REGION Network 26: Head status
   RUNG wire#powerrail
      Contact( "AlwaysTRUE" )
      wire#w1
      I_Contact( #OUTPUT_xFireON )
      Move(in := 1, out1 => #tHMR.dHeadStatus)
   END_RUNG
   RUNG wire#w1
      Contact( #OUTPUT_xFireON )
      Move(in := 3, out1 => #tHMR.dHeadStatus)
   END_RUNG
   // the same network as SCL:
   IF "AlwaysTRUE" AND NOT #OUTPUT_xFireON THEN #tHMR.dHeadStatus := 1; END_IF;
   IF "AlwaysTRUE" AND #OUTPUT_xFireON THEN #tHMR.dHeadStatus := 3; END_IF;
END_REGION

REGION Network 27: Head#x reset head usage counter {x|x|x|x|O}
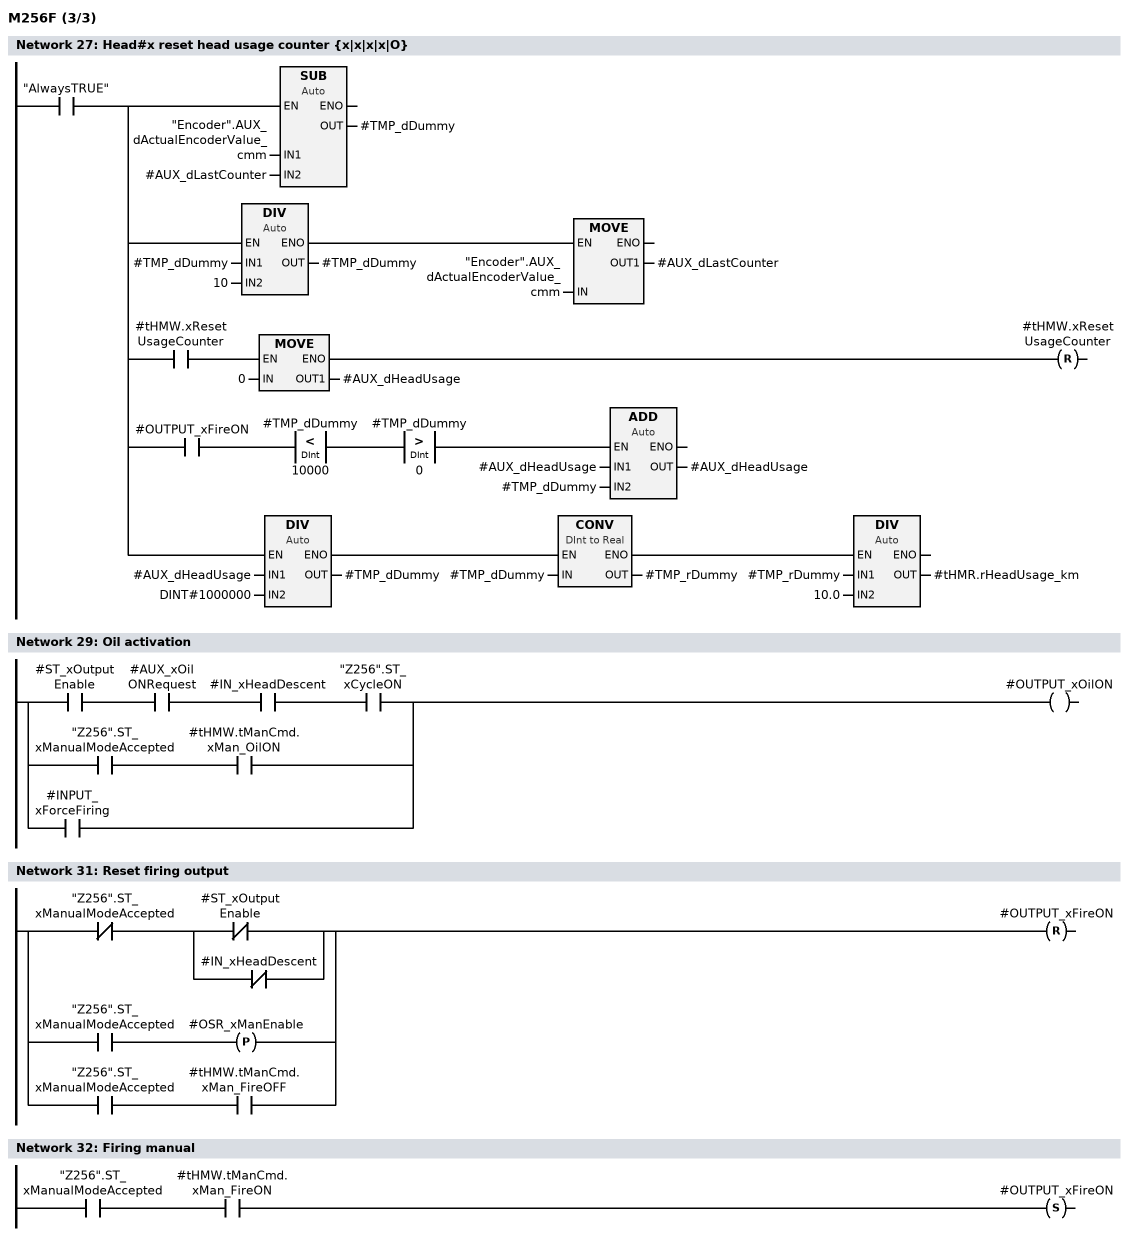
   RUNG wire#powerrail
      Contact( "AlwaysTRUE" )
      wire#w1
      Sub(in1 := "Encoder".AUX_dActualEncoderValue_cmm, in2 := #AUX_dLastCounter, out => #TMP_dDummy)
   END_RUNG
   RUNG wire#w1
      Div(in1 := #TMP_dDummy, in2 := 10, out => #TMP_dDummy)
      Move(in := "Encoder".AUX_dActualEncoderValue_cmm, out1 => #AUX_dLastCounter)
   END_RUNG
   RUNG wire#w1
      Contact( #tHMW.xResetUsageCounter )
      Move(in := 0, out1 => #AUX_dHeadUsage)
      R_Coil( #tHMW.xResetUsageCounter )
   END_RUNG
   RUNG wire#w1
      Contact( #OUTPUT_xFireON )
      { S7_Templates := "SrcType := DInt" } LT_Contact(in1 := #TMP_dDummy, in2 := 10000)
      { S7_Templates := "SrcType := DInt" } GT_Contact(in1 := #TMP_dDummy, in2 := 0)
      Add(in1 := #AUX_dHeadUsage, in2 := #TMP_dDummy, out => #AUX_dHeadUsage)
   END_RUNG
   RUNG wire#w1
      Div(in1 := #AUX_dHeadUsage, in2 := DINT#1000000, out => #TMP_dDummy)
      { S7_Templates := "[SrcType := DInt, DestType := Real]" } Convert(in := #TMP_dDummy, out => #TMP_rDummy)
      Div(in1 := #TMP_rDummy, in2 := 10.0, out => #tHMR.rHeadUsage_km)
   END_RUNG
   // the same network as SCL:
   IF "AlwaysTRUE" THEN
       #TMP_dDummy := "Encoder".AUX_dActualEncoderValue_cmm - #AUX_dLastCounter;
       #TMP_dDummy := #TMP_dDummy / 10;
       #AUX_dLastCounter := "Encoder".AUX_dActualEncoderValue_cmm;
   END_IF;
   IF "AlwaysTRUE" AND #tHMW.xResetUsageCounter THEN
       #AUX_dHeadUsage := 0;
       #tHMW.xResetUsageCounter := FALSE;
   END_IF;
   IF "AlwaysTRUE" AND #OUTPUT_xFireON AND (#TMP_dDummy < 10000) AND (#TMP_dDummy > 0) THEN
       #AUX_dHeadUsage := #AUX_dHeadUsage + #TMP_dDummy;
   END_IF;
   IF "AlwaysTRUE" THEN
       #TMP_dDummy := #AUX_dHeadUsage / DINT#1000000;
       #TMP_rDummy := DINT_TO_REAL(#TMP_dDummy);
       #tHMR.rHeadUsage_km := #TMP_rDummy / 10.0;
   END_IF;
END_REGION

REGION Network 28: ####_OUTPUT_####
END_REGION

REGION Network 29: Oil activation
   RUNG wire#powerrail
      Contact( #ST_xOutputEnable )
      Contact( #AUX_xOilONRequest )
      Contact( #IN_xHeadDescent )
      Contact( "Z256".ST_xCycleON )
      wire#w1
      Coil( #OUTPUT_xOilON )
   END_RUNG
   RUNG wire#powerrail
      Contact( "Z256".ST_xManualModeAccepted )
      Contact( #tHMW.tManCmd.xMan_OilON )
   END_RUNG wire#w1
   RUNG wire#powerrail
      Contact( #INPUT_xForceFiring )
   END_RUNG wire#w1
   // the same network as SCL:
   #OUTPUT_xOilON := (#ST_xOutputEnable AND #AUX_xOilONRequest AND #IN_xHeadDescent AND "Z256".ST_xCycleON) OR ("Z256".ST_xManualModeAccepted AND #tHMW.tManCmd.xMan_OilON) OR #INPUT_xForceFiring;
END_REGION

REGION Network 30 (SCL): Pressure to heads and display
   #TMP_rDummy := DINT_TO_REAL("CONST_dPressureMax_Unit"-"CONST_dPressureMin_Unit")/ DINT_TO_REAL("CONST_dPressureMax_MN"-"CONST_dPressureMin_MN");
   #TMP_dDummy :=#tHMW.dHeadPressure_mN-"CONST_dPressureMin_MN";
   #OUTPUT_iPressuremA := REAL_TO_INT(#TMP_rDummy *  DINT_TO_REAL(#TMP_dDummy))+DINT_TO_INT("CONST_dPressureMin_Unit");

   IF "CM_IDEV_FromMainLine".xQLTplate THEN
       #OUTPUT_iPressuremA := #OUTPUT_iPressuremA / 100 * DINT_TO_INT("Z256_hmi".tHMW.dPressureScalerOnSample_perc);
   END_IF;
END_REGION

REGION Network 31: Reset firing output
   RUNG wire#powerrail
      I_Contact( "Z256".ST_xManualModeAccepted )
      wire#w1
      I_Contact( #ST_xOutputEnable )
      wire#w2
      R_Coil( #OUTPUT_xFireON )
   END_RUNG
   RUNG wire#w1
      I_Contact( #IN_xHeadDescent )
   END_RUNG wire#w2
   RUNG wire#powerrail
      Contact( "Z256".ST_xManualModeAccepted )
      P_Trig( #OSR_xManEnable )
   END_RUNG wire#w2
   RUNG wire#powerrail
      Contact( "Z256".ST_xManualModeAccepted )
      Contact( #tHMW.tManCmd.xMan_FireOFF )
   END_RUNG wire#w2
   // the same network as SCL:
   #_w1 := "Z256".ST_xManualModeAccepted AND NOT #OSR_xManEnable;   // rising edge
   #OSR_xManEnable := "Z256".ST_xManualModeAccepted;
   IF (NOT "Z256".ST_xManualModeAccepted AND (NOT #ST_xOutputEnable OR NOT #IN_xHeadDescent)) OR #_w1 OR ("Z256".ST_xManualModeAccepted AND #tHMW.tManCmd.xMan_FireOFF) THEN
       #OUTPUT_xFireON := FALSE;
   END_IF;
END_REGION

REGION Network 32: Firing manual
   RUNG wire#powerrail
      Contact( "Z256".ST_xManualModeAccepted )
      Contact( #tHMW.tManCmd.xMan_FireON )
      S_Coil( #OUTPUT_xFireON )
   END_RUNG
   // the same network as SCL:
   IF "Z256".ST_xManualModeAccepted AND #tHMW.tManCmd.xMan_FireON THEN #OUTPUT_xFireON := TRUE; END_IF;
END_REGION
END_FUNCTION_BLOCK

FUNCTION_BLOCK "M256M"   // FB101, LAD
{ S7_Optimized_Access := 'TRUE' }
VERSION : 0.1
   VAR_INPUT
      IN_tConnectionData : "UDT_MB_ConnData";   // IP and connection ID
      IN_dHeadCycleIndex : DInt;   // Number of head cycle (Actual head-1)
      IN_xST_AllHeadStoppingFaults : Bool;   // Cumulative head alarm
      IN_ST_xAllHeadInitialized : Bool;   // All head initialized
      IN_ST_xAllHeadPositioned : Bool;   // All head positioned
      IN_ST_xAllHeadReferred : Bool;   // All head referred
   END_VAR
   VAR
      ST_xHeadInitialized : Bool;   // Head #x initialized
      ST_xHeadReferredSwitch : Bool;   // Head #x referred
      ST_xHeadPositioned : Bool;   // Head #x positioned
      ST_xOutputEnable : Bool;   // Head #x output enable
      ST_xPhaseInProgress : Bool;   // Head #x phases in progress
      ST_xStoppingFaults : Bool;   // Head #x in stopping fault
      ST_xWarnings : Bool;   // Head #x in warning
      ST_xMovementInProgress : Bool;   // Head #x in movement
      ST_xFaults : Bool;   // Head #x in faults
      ST_xHeadVirtualCollision : Bool;   // Head #x virtual collision
      ST_xHeadIPAvail : Bool;   // Head #x is IP linked
      ST_xBrakeReleaseRequest : Bool;   // Head #x brake release requested
      ST_xConditionOKforPowerON : Bool;   // Head #x power on condition
      OSR_xAllHeadReferred : Bool;   // OSR all hed referred
      OSR_xDriveEnable : Bool;   // OSR drive enable
      OSR_xBrakeReleaseSB : Bool;   // OS Brake release
      OS_xBrakeReleaseSB : Bool;   // OS Brake release
      OS_xBrakeRelease : Bool;   // OS Brake release
      OS_xBrakeEngage : Bool;   // OS Brake engaged
      ON_xMotorMBReset : Bool;   // ON Modbus motor reset
      OSN_xMotorMBReset : Bool;   // OSN Modbus motor reset
      INPUT_xOverstroke : Bool;   // Head #x Carriage overstroke
      INPUT_xBrakeRelease : Bool;   // Head #x Brake release button
      INPUT_xCarriageOverload : Bool;   // Head #x Carriage overload
      PH_xHeadInit : Bool;   // Head #x initialization in progress
      PH_xHeadEndInit : Bool;   // Head #x end initialization in progress
      PH_xHeadHomeSwitch : Bool;   // Head #x home in progress to switch
      PH_xHeadEndHomeSwitch : Bool;   // Head #x end home in progress to switch
      PH_xHeadPositioning : Bool;   // Head #x positioning in progress
      PH_xHeadEndPositioning : Bool;   // Head #x end positioning in progress
      AUX_tModbusTCP : TCP_MB_FC8_Req;   // Modbus data
      AUX_xPosCadencer : Bool;   // Cadencer head #x - Positioning allowed
      AUX_dHeadRequestPosition_cmm : DInt;   // Head #x request position [mm/100]
      AUX_dHeadActualPosition_cmm : DInt;   // Head #x actual position [mm/100]
      AUX_rDistanceSwitchTo0 : Real;   // Head #x distance 0 encoder to cam
      AUX_dHeadActSpeed : DInt;   // Head #x actual speed
      AUX_dActualDownloadPar : DInt;   // Head #x actual parameter in download
      AUX_xHomeCadencer : Bool;   // Cadencer head #x - Home position allowed
      AUX_tmDriveReadyRetainTimer : IEC_TIMER;   // Drive ready retain timer
      AUX_tmHeadPositioningTimeout : IEC_TIMER;   // Positioning timeout timer
      AUX_tmHeadHomingTimeout : IEC_TIMER;   // Homing timeout timer
      AUX_tmOFFComOK : IEC_TIMER;   // Head communication OK retained
      AUX_tmOFFEnablePositioningAfterHome : IEC_TIMER;   // Wait drive positioning after homing
      AUX_tmOFFDriveEnable : IEC_TIMER;   // Wait drive enable
      AUX_tmOFFReadCamOffsetAfterHome : IEC_TIMER;   // Retained read cam offset after homing
      AUX_tmHeadInitTimeout : IEC_TIMER;   // Initialization timeout timer
      Axis_Ref : "ILx2T_Ref";
      ILx2_ModbusTCP_Data_Instance : "ILx2_ModbusTCP_Data_1500";
      ILx2T_Control_Instance : "ILx2T_Control";
      ILx2T_Homing_Instance : "ILx2T_Homing";
      ILx2T_Jog_Instance : "ILx2T_Jog";
      ILx2T_ProfilePosition_Instance : "ILx2T_ProfilePosition";
      ILx2T_ProfileVelocity_Instance : "ILx2T_ProfileVelocity";
      ILx2T_Parameter_Read_Write_Instance_Pos : "ILx2T_Parameter_Read_Write";
      ILx2T_Parameter_Read_Write_Instance_Cam : "ILx2T_Parameter_Read_Write";
      ILx2T_Parameter_Read_Write_Instance_Speed : "ILx2T_Parameter_Read_Write";
      ILx2T_Parameter_Read_Write_Instance : "ILx2T_Parameter_Read_Write";
   END_VAR
   VAR RETAIN
      tHMR : Struct   // {[Unit][Scada unit][Low limit][High limit][Access]}
         iCodeAlarm : Int;
         dHeadActualPositions_cmm : DInt;   // Head#x head actual position [mm/100] {mm/100|mm|x|x|O} / Head #x head actual position [mm/100] {mm/100|mm|x|x|O}
         dHeadHomePositions_cmm : DInt;   // Head#x home position [mm/100] {mm/100|mm|x|x|O} / Head #x home position [mm/100] {mm/100|mm|x|x|O}
         rgdHeadMoveStatus : DInt;   // Head#x move status (1=Not Initialized 2=Not referred 3=Not positioned 4=Positioned 5=Positioning 6=Virtual collision 7=Anomaly) {x|x|x|x|O} / Head #x move status (1=Not Initialized 2=Not referred 3=Not positioned 4=Positioned 5=Positioning 6=Virtual collision 7=Anomaly) {x|x|x|x|O}
         tManCmd : Struct
            xMan_JogForwardFdbk : Bool;   // Head#x manual jog forward fdbk {x|x|x|x|O} / Head #x manual jog forward fdbk {x|x|x|x|O}
            xMan_JogBackwardFdbk : Bool;   // Head#x manual jog backward fdbk {x|x|x|x|O} / Head #x manual jog backward fdbk {x|x|x|x|O}
         END_STRUCT;
      END_STRUCT;
      tHMW : Struct   // {[Unit][Scada unit][Low limit][High limit][Access]}
         xBrakeRealeaseHeads : Bool := FALSE;   // Force the brake release of the head {x|x|x|x|M}
         xBrakeEngageHeads : Bool := FALSE;   // Force the brake engaged of the head {x|x|x|x|M}
         xUpdateHomeHead : Bool;   // Update home position head#x {x|x|x|x|M} / Update home position Head #x {x|x|x|x|M}
         dHeadHomePositions_cmm : DInt;   // Head#x home position [mm/100] {mm/100|mm|-2500|2500|M} / Head #x home position [mm/100] {mm/100|mm|-2500|2500|M}
         tManCmd : Struct
            xMan_JogBackward : Bool;   // Head #x manual jog backward {x|x|x|x|O}
            xMan_JogForward : Bool;   // Head #x manual jog forward {x|x|x|x|O}
         END_STRUCT;
      END_STRUCT;
   END_VAR
   VAR
      tALM : Struct
         tW : Struct
            x0 : Bool;
            x1 : Bool;
            x2 : Bool;
            x3 : Bool;
            x4 : Bool;
            x5 : Bool;
            x6 : Bool;
            x7 : Bool;
            x8 : Bool;
            x9 : Bool;
            x10 : Bool;
            x11 : Bool;
            x12 : Bool;
            x13 : Bool;
            x14 : Bool;
            x15 : Bool;
            x16 : Bool;
            x17 : Bool;
            x18 : Bool;
            x19 : Bool;
            x20 : Bool;
            x21 : Bool;
            x22 : Bool;
            x23 : Bool;
            x24 : Bool;
            x25 : Bool;
            x26 : Bool;
            x27 : Bool;
            x28 : Bool;
            x29 : Bool;
            x30 : Bool;
            x31 : Bool;
         END_STRUCT;
         tS : Struct
            x0 : Bool;   // Head#x Initialization timeout / Head #x Initialization timeout
            x1 : Bool;   // Head#x homing timeout / Head #x homing timeout
            x2 : Bool;   // Head#x positioning timeout / Head #x positioning timeout
            x3 : Bool;   // Head#x carriage overload / Head #x carriage overload
            x4 : Bool;   // Head#x drive error / Head #x drive error
            x5 : Bool;   // Head#x missing ethernet IP connection / Head #x missing ethernet IP connection
            x6 : Bool;   // Head op.side overstroke
            x7 : Bool;   // Head oppo.op.side overstroke
            x8 : Bool;   // Head #x overstroke
            x9 : Bool;
            x10 : Bool;
            x11 : Bool;
            x12 : Bool;
            x13 : Bool;
            x14 : Bool;
            x15 : Bool;
            x16 : Bool;
            x17 : Bool;
            x18 : Bool;
            x19 : Bool;
            x20 : Bool;
            x21 : Bool;
            x22 : Bool;
            x23 : Bool;
            x24 : Bool;
            x25 : Bool;
            x26 : Bool;
            x27 : Bool;
            x28 : Bool;
            x29 : Bool;
            x30 : Bool;
            x31 : Bool;
         END_STRUCT;
         tF : Struct
            x0 : Bool;
            x1 : Bool;
            x2 : Bool;
            x3 : Bool;
            x4 : Bool;
            x5 : Bool;
            x6 : Bool;
            x7 : Bool;
            x8 : Bool;
            x9 : Bool;
            x10 : Bool;
            x11 : Bool;
            x12 : Bool;
            x13 : Bool;
            x14 : Bool;
            x15 : Bool;
            x16 : Bool;
            x17 : Bool;
            x18 : Bool;
            x19 : Bool;
            x20 : Bool;
            x21 : Bool;
            x22 : Bool;
            x23 : Bool;
            x24 : Bool;
            x25 : Bool;
            x26 : Bool;
            x27 : Bool;
            x28 : Bool;
            x29 : Bool;
            x30 : Bool;
            x31 : Bool;
         END_STRUCT;
      END_STRUCT;
   END_VAR
   VAR_TEMP
      TMP_rDummy : Real;
      TMP_dwDummy : DWord;
      TMP_dDummy : DInt;
      TMP_dPosition : DInt;
      TMP_dIndex2Nd : DInt;
      TMP_xWriteDoneOS : Bool;
      TMP_xRead : Bool;
      TMP_xMotorOFF : Bool;
   END_VAR
   VAR_TEMP   // added for the SCL form of the ladder/FBD networks
      _w1 : Bool;
      _w2 : Bool;
   END_VAR
   // ILx2T_Homing_Instance.i_diHMsrchdisusr := 0;
BEGIN

REGION Network 1: ####_COSTANTS_####
END_REGION

REGION Network 2: ####_ALARMS_####
END_REGION

REGION Network 3: Reset faults
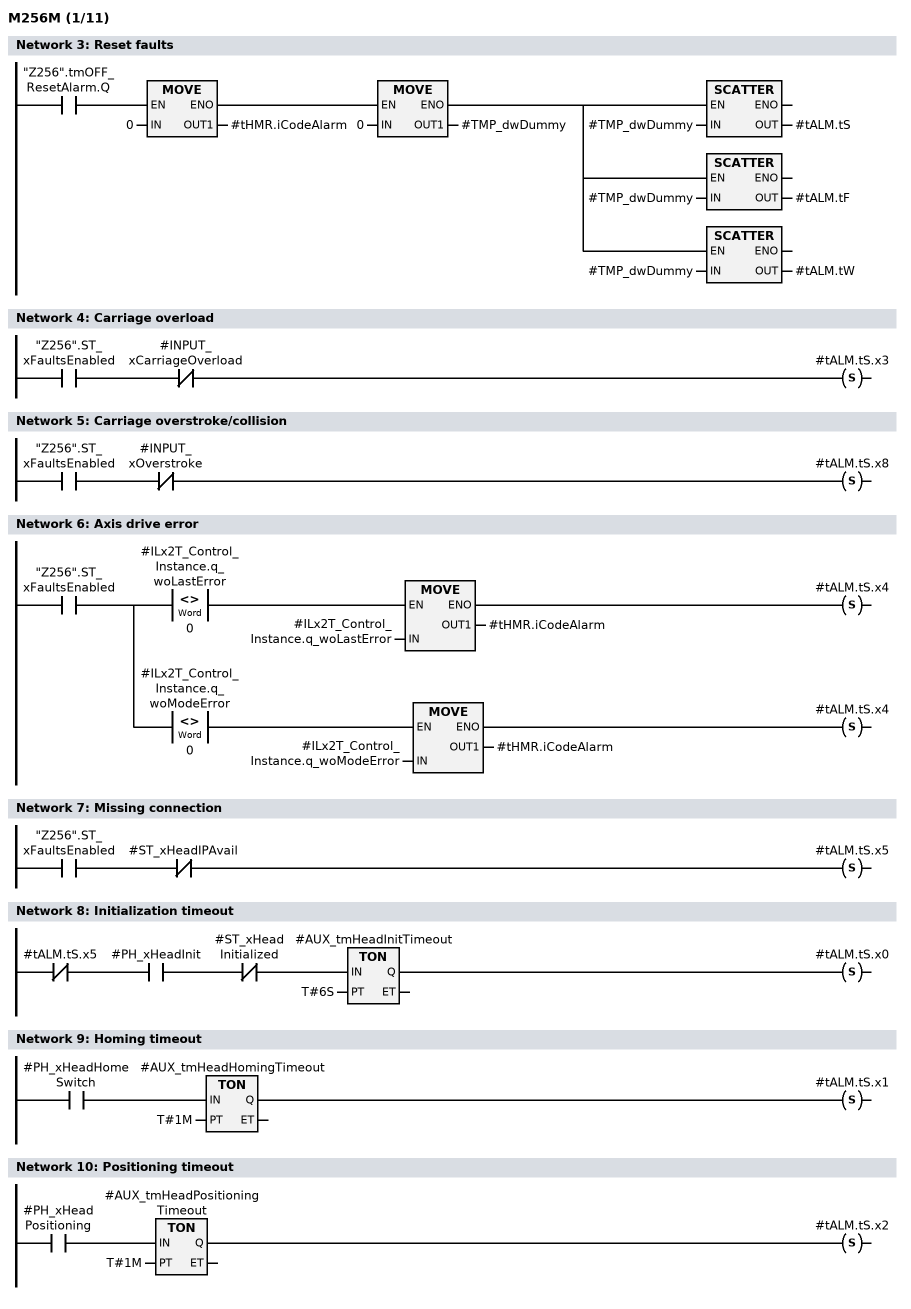
   IF "Z256".tmOFF_ResetAlarm.Q THEN
       #tHMR.iCodeAlarm := 0;
       #TMP_dwDummy := 0;
   END_IF;
   #_w1 := "Z256".tmOFF_ResetAlarm.Q;
   IF #_w1 THEN
       SCATTER(IN := #TMP_dwDummy, OUT => #tALM.tS);
       SCATTER(IN := #TMP_dwDummy, OUT => #tALM.tF);
       SCATTER(IN := #TMP_dwDummy, OUT => #tALM.tW);
   END_IF;
END_REGION

REGION Network 4: Carriage overload
   RUNG wire#powerrail
      Contact( "Z256".ST_xFaultsEnabled )
      I_Contact( #INPUT_xCarriageOverload )
      S_Coil( #tALM.tS.x3 )
   END_RUNG
   // the same network as SCL:
   IF "Z256".ST_xFaultsEnabled AND NOT #INPUT_xCarriageOverload THEN #tALM.tS.x3 := TRUE; END_IF;
END_REGION

REGION Network 5: Carriage overstroke/collision
   RUNG wire#powerrail
      Contact( "Z256".ST_xFaultsEnabled )
      I_Contact( #INPUT_xOverstroke )
      S_Coil( #tALM.tS.x8 )
   END_RUNG
   // the same network as SCL:
   IF "Z256".ST_xFaultsEnabled AND NOT #INPUT_xOverstroke THEN #tALM.tS.x8 := TRUE; END_IF;
END_REGION

REGION Network 6: Axis drive error
   RUNG wire#powerrail
      Contact( "Z256".ST_xFaultsEnabled )
      wire#w1
      { S7_Templates := "SrcType := Word" } NE_Contact(in1 := #ILx2T_Control_Instance.q_woLastError, in2 := 0)
      Move(in := #ILx2T_Control_Instance.q_woLastError, out1 => #tHMR.iCodeAlarm)
      S_Coil( #tALM.tS.x4 )
   END_RUNG
   RUNG wire#w1
      { S7_Templates := "SrcType := Word" } NE_Contact(in1 := #ILx2T_Control_Instance.q_woModeError, in2 := 0)
      Move(in := #ILx2T_Control_Instance.q_woModeError, out1 => #tHMR.iCodeAlarm)
      S_Coil( #tALM.tS.x4 )
   END_RUNG
   // the same network as SCL:
   IF "Z256".ST_xFaultsEnabled AND (#ILx2T_Control_Instance.q_woLastError <> 0) THEN
       #tHMR.iCodeAlarm := #ILx2T_Control_Instance.q_woLastError;
       #tALM.tS.x4 := TRUE;
   END_IF;
   IF "Z256".ST_xFaultsEnabled AND (#ILx2T_Control_Instance.q_woModeError <> 0) THEN
       #tHMR.iCodeAlarm := #ILx2T_Control_Instance.q_woModeError;
       #tALM.tS.x4 := TRUE;
   END_IF;
END_REGION

REGION Network 7: Missing connection
   RUNG wire#powerrail
      Contact( "Z256".ST_xFaultsEnabled )
      I_Contact( #ST_xHeadIPAvail )
      S_Coil( #tALM.tS.x5 )
   END_RUNG
   // the same network as SCL:
   IF "Z256".ST_xFaultsEnabled AND NOT #ST_xHeadIPAvail THEN #tALM.tS.x5 := TRUE; END_IF;
END_REGION

REGION Network 8: Initialization timeout
   #AUX_tmHeadInitTimeout.TON(IN := NOT #tALM.tS.x5 AND #PH_xHeadInit AND NOT #ST_xHeadInitialized, PT := T#6S);
   IF #AUX_tmHeadInitTimeout.Q THEN #tALM.tS.x0 := TRUE; END_IF;
END_REGION

REGION Network 9: Homing timeout
   #AUX_tmHeadHomingTimeout.TON(IN := #PH_xHeadHomeSwitch, PT := T#1M);
   IF #AUX_tmHeadHomingTimeout.Q THEN #tALM.tS.x1 := TRUE; END_IF;
END_REGION

REGION Network 10: Positioning timeout
   #AUX_tmHeadPositioningTimeout.TON(IN := #PH_xHeadPositioning, PT := T#1M);
   IF #AUX_tmHeadPositioningTimeout.Q THEN #tALM.tS.x2 := TRUE; END_IF;
END_REGION

REGION Network 11 (SCL): Cumulative of warning active
   #ST_xWarnings := 0;

   GATHER(IN:= #tALM.tW,
          OUT=>#TMP_dwDummy);

   IF #TMP_dwDummy <> 0 THEN
       #ST_xWarnings := 1;
   END_IF;
END_REGION

REGION Network 12 (SCL): Cumulative of stopping faults active
   #ST_xStoppingFaults := 0;
   GATHER(IN := #tALM.tS,
          OUT => #TMP_dwDummy);

   IF #TMP_dwDummy <> 0 THEN
       #ST_xStoppingFaults := 1;
   END_IF;
END_REGION

REGION Network 13 (SCL): Cumulative of faults active
   #ST_xFaults := 0;
   GATHER(IN := #tALM.tF,
          OUT => #TMP_dwDummy);

   IF #TMP_dwDummy <> 0 THEN
       #ST_xFaults := 1;
   END_IF;
END_REGION

REGION Network 14: #####_HMI LOGICS_#####
END_REGION

REGION Network 15: OS Brake release
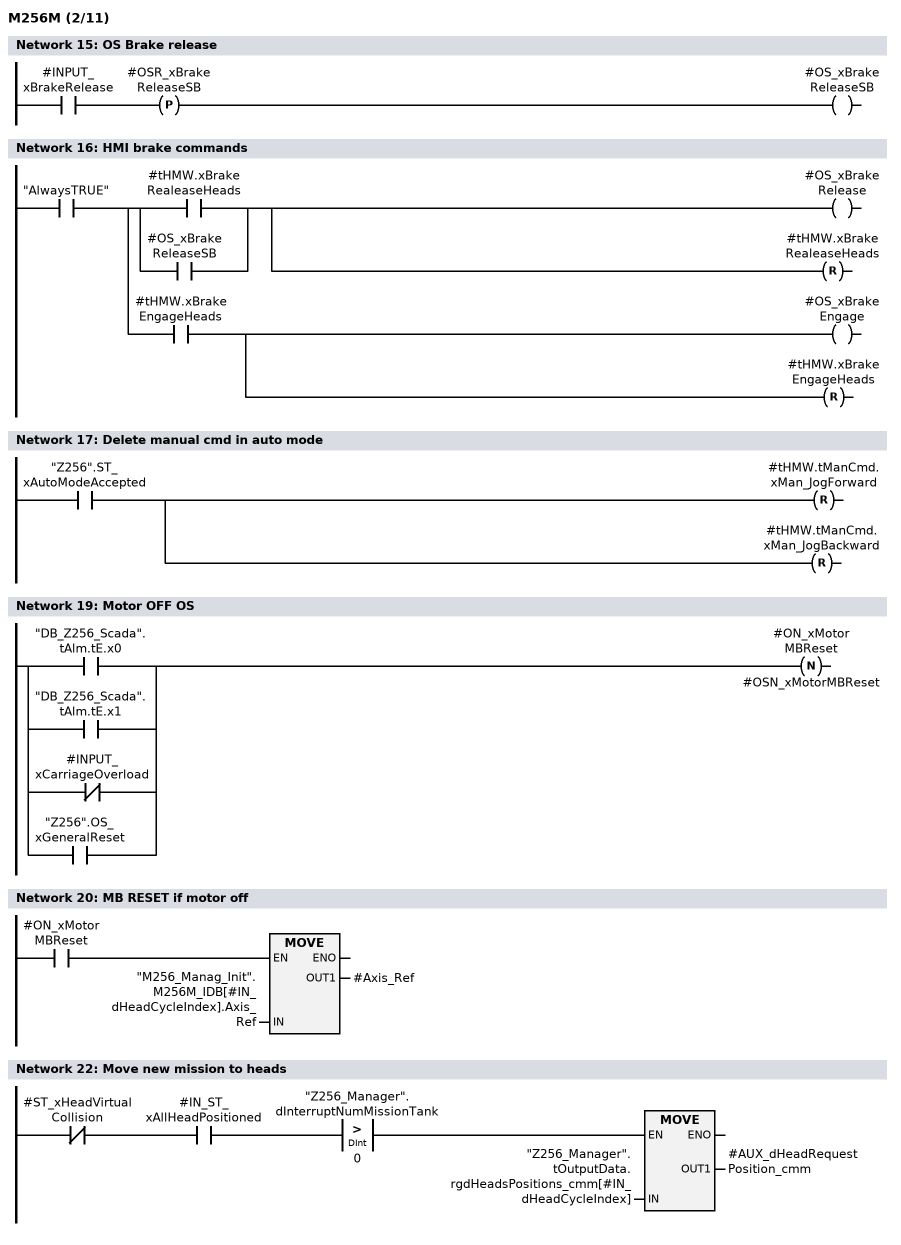
   RUNG wire#powerrail
      Contact( #INPUT_xBrakeRelease )
      P_Trig( #OSR_xBrakeReleaseSB )
      Coil( #OS_xBrakeReleaseSB )
   END_RUNG
   // the same network as SCL:
   #_w1 := #INPUT_xBrakeRelease AND NOT #OSR_xBrakeReleaseSB;   // rising edge
   #OSR_xBrakeReleaseSB := #INPUT_xBrakeRelease;
   #OS_xBrakeReleaseSB := #_w1;
END_REGION

REGION Network 16: HMI brake commands
   RUNG wire#powerrail
      Contact( "AlwaysTRUE" )
      wire#w1
      Contact( #tHMW.xBrakeRealeaseHeads )
      wire#w2
      Coil( #OS_xBrakeRelease )
   END_RUNG
   RUNG wire#w1
      Contact( #OS_xBrakeReleaseSB )
   END_RUNG wire#w2
   RUNG wire#w2
      R_Coil( #tHMW.xBrakeRealeaseHeads )
   END_RUNG
   RUNG wire#w1
      Contact( #tHMW.xBrakeEngageHeads )
      wire#w3
      Coil( #OS_xBrakeEngage )
   END_RUNG
   RUNG wire#w3
      R_Coil( #tHMW.xBrakeEngageHeads )
   END_RUNG
   // the same network as SCL:
   #OS_xBrakeRelease := "AlwaysTRUE" AND (#tHMW.xBrakeRealeaseHeads OR #OS_xBrakeReleaseSB);
   IF #OS_xBrakeRelease THEN #tHMW.xBrakeRealeaseHeads := FALSE; END_IF;
   #OS_xBrakeEngage := "AlwaysTRUE" AND #tHMW.xBrakeEngageHeads;
   IF #OS_xBrakeEngage THEN #tHMW.xBrakeEngageHeads := FALSE; END_IF;
END_REGION

REGION Network 17: Delete manual cmd in auto mode
   RUNG wire#powerrail
      Contact( "Z256".ST_xAutoModeAccepted )
      wire#w1
      R_Coil( #tHMW.tManCmd.xMan_JogForward )
   END_RUNG
   RUNG wire#w1
      R_Coil( #tHMW.tManCmd.xMan_JogBackward )
   END_RUNG
   // the same network as SCL:
   IF "Z256".ST_xAutoModeAccepted THEN
       #tHMW.tManCmd.xMan_JogForward := FALSE;
       #tHMW.tManCmd.xMan_JogBackward := FALSE;
   END_IF;
END_REGION

REGION Network 18: #####_ILA2 MANAGEMENT_#####
END_REGION

REGION Network 19: Motor OFF OS
   #_w1 := "DB_Z256_Scada".tAlm.tE.x0 OR "DB_Z256_Scada".tAlm.tE.x1 OR NOT #INPUT_xCarriageOverload OR "Z256".OS_xGeneralReset;
   #ON_xMotorMBReset := NOT #_w1 AND #OSN_xMotorMBReset;   // falling edge
   #OSN_xMotorMBReset := #_w1;
END_REGION

REGION Network 20: MB RESET if motor off
   RUNG wire#powerrail
      Contact( #ON_xMotorMBReset )
      Move(in := "M256_Manag_Init".M256M_IDB[#IN_dHeadCycleIndex].Axis_Ref, out1 => #Axis_Ref)
   END_RUNG
   // the same network as SCL:
   IF #ON_xMotorMBReset THEN #Axis_Ref := "M256_Manag_Init".M256M_IDB[#IN_dHeadCycleIndex].Axis_Ref; END_IF;
END_REGION

REGION Network 21 (SCL): MB RESET if motor off
   IF #ON_xMotorMBReset THEN
       #ILx2_ModbusTCP_Data_Instance.Com_OK := 0;
       #ILx2_ModbusTCP_Data_Instance.diErrorCounter_DPL_Read := 0;
       #ILx2_ModbusTCP_Data_Instance.diErrorCounter_DPL_Write := 0;
       #ILx2_ModbusTCP_Data_Instance.diErrorCounter_Para_Read := 0;
       #ILx2_ModbusTCP_Data_Instance.diErrorCounter_Para_Write := 0;
       #ILx2_ModbusTCP_Data_Instance.Index := 0;
       #ILx2_ModbusTCP_Data_Instance.inIndex := 0;
       #ILx2_ModbusTCP_Data_Instance.Error := 0;
       #ILx2_ModbusTCP_Data_Instance.xErrorReadDPL := 0;
       #ILx2_ModbusTCP_Data_Instance.xErrorWriteDPL := 0;
       #ILx2_ModbusTCP_Data_Instance.xErrorReadParameter := 0;
       #ILx2_ModbusTCP_Data_Instance.xErrorWriteParameter := 0;
       #ILx2_ModbusTCP_Data_Instance.xNodeGuardInitOK := 0;
       #ILx2_ModbusTCP_Data_Instance.Index := 0;
       #ILx2_ModbusTCP_Data_Instance.inIndex := 0;
       #ILx2_ModbusTCP_Data_Instance.inNodeGuardTime := 0;
       #ILx2_ModbusTCP_Data_Instance.iState_Read_DPL := 0;
       #ILx2_ModbusTCP_Data_Instance.iState_Write_DPL := 0;
       #ILx2_ModbusTCP_Data_Instance.iState_Read_Para := 0;
       #ILx2_ModbusTCP_Data_Instance.iState_Write_Para := 0;
       #ILx2_ModbusTCP_Data_Instance.iStateTimeReadDPL := 0;
       #ILx2_ModbusTCP_Data_Instance.iStateTimeWriteDPL := 0;
       #ILx2_ModbusTCP_Data_Instance.ParaRead_Value := 0;
       #ILx2_ModbusTCP_Data_Instance.ParaWrite_Value := 0;
       #ILx2_ModbusTCP_Data_Instance.ReadData_DPL := "M256_Manag_Init".M256M_IDB[#IN_dHeadCycleIndex].ILx2_ModbusTCP_Data_Instance.ReadData_DPL;
       #ILx2_ModbusTCP_Data_Instance.WriteData_DPL := "M256_Manag_Init".M256M_IDB[#IN_dHeadCycleIndex].ILx2_ModbusTCP_Data_Instance.WriteData_DPL;
       #ILx2_ModbusTCP_Data_Instance.stCONNECT_DPL_Read := "M256_Manag_Init".M256M_IDB[#IN_dHeadCycleIndex].ILx2_ModbusTCP_Data_Instance.stCONNECT_DPL_Read;
       #ILx2_ModbusTCP_Data_Instance.stCONNECT_DPL_Write := "M256_Manag_Init".M256M_IDB[#IN_dHeadCycleIndex].ILx2_ModbusTCP_Data_Instance.stCONNECT_DPL_Write;
       #ILx2_ModbusTCP_Data_Instance.stCONNECT_Parameter_Read := "M256_Manag_Init".M256M_IDB[#IN_dHeadCycleIndex].ILx2_ModbusTCP_Data_Instance.stCONNECT_Parameter_Read;
       #ILx2_ModbusTCP_Data_Instance.stCONNECT_Parameter_Write := "M256_Manag_Init".M256M_IDB[#IN_dHeadCycleIndex].ILx2_ModbusTCP_Data_Instance.stCONNECT_Parameter_Write;
       #ILx2_ModbusTCP_Data_Instance.xNodeGuardInitOK := 0;
   END_IF;
END_REGION

REGION Network 22: Move new mission to heads
   RUNG wire#powerrail
      I_Contact( #ST_xHeadVirtualCollision )
      Contact( #IN_ST_xAllHeadPositioned )
      { S7_Templates := "SrcType := DInt" } GT_Contact(in1 := "Z256_Manager".dInterruptNumMissionTank, in2 := 0)
      Move(in := "Z256_Manager".tOutputData.rgdHeadsPositions_cmm[#IN_dHeadCycleIndex], out1 => #AUX_dHeadRequestPosition_cmm)
   END_RUNG
   // the same network as SCL:
   IF NOT #ST_xHeadVirtualCollision AND #IN_ST_xAllHeadPositioned AND ("Z256_Manager".dInterruptNumMissionTank > 0) THEN
       #AUX_dHeadRequestPosition_cmm := "Z256_Manager".tOutputData.rgdHeadsPositions_cmm[#IN_dHeadCycleIndex];
   END_IF;
END_REGION

REGION Network 23: MB Connection
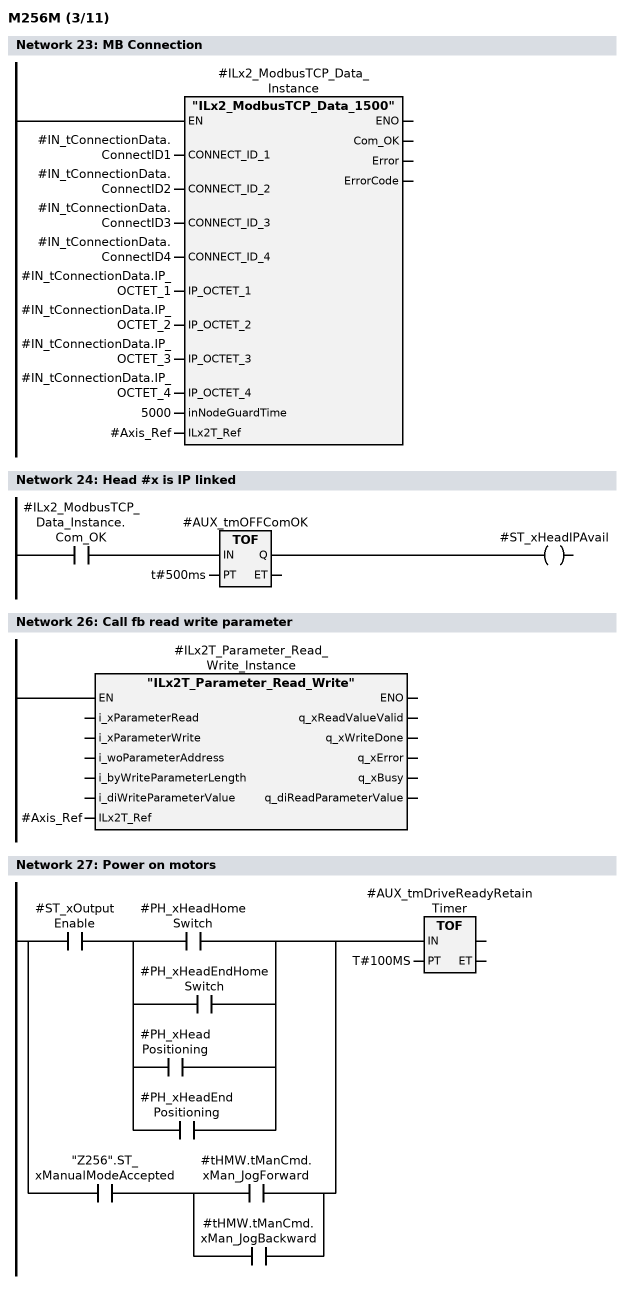
   RUNG wire#powerrail
      #ILx2_ModbusTCP_Data_Instance(CONNECT_ID_1 := #IN_tConnectionData.ConnectID1, CONNECT_ID_2 := #IN_tConnectionData.ConnectID2, CONNECT_ID_3 := #IN_tConnectionData.ConnectID3, CONNECT_ID_4 := #IN_tConnectionData.ConnectID4, IP_OCTET_1 := #IN_tConnectionData.IP_OCTET_1, IP_OCTET_2 := #IN_tConnectionData.IP_OCTET_2, IP_OCTET_3 := #IN_tConnectionData.IP_OCTET_3, IP_OCTET_4 := #IN_tConnectionData.IP_OCTET_4, inNodeGuardTime := 5000, ILx2T_Ref := #Axis_Ref, Com_OK =>, Error =>, ErrorCode =>)
   END_RUNG
   // the same network as SCL:
   #ILx2_ModbusTCP_Data_Instance(CONNECT_ID_1 := #IN_tConnectionData.ConnectID1,   // "ILx2_ModbusTCP_Data_1500"
                           CONNECT_ID_2 := #IN_tConnectionData.ConnectID2,
                           CONNECT_ID_3 := #IN_tConnectionData.ConnectID3,
                           CONNECT_ID_4 := #IN_tConnectionData.ConnectID4,
                           IP_OCTET_1 := #IN_tConnectionData.IP_OCTET_1,
                           IP_OCTET_2 := #IN_tConnectionData.IP_OCTET_2,
                           IP_OCTET_3 := #IN_tConnectionData.IP_OCTET_3,
                           IP_OCTET_4 := #IN_tConnectionData.IP_OCTET_4,
                           inNodeGuardTime := 5000,
                           ILx2T_Ref := #Axis_Ref);
END_REGION

REGION Network 24: Head #x is IP linked
   #AUX_tmOFFComOK.TOF(IN := #ILx2_ModbusTCP_Data_Instance.Com_OK, PT := t#500ms);
   #ST_xHeadIPAvail := #AUX_tmOFFComOK.Q;
END_REGION

REGION Network 25 (SCL): Head Init - Download parameters
   //THIS SUBROUTINE WILL INITIALIZE ALL THE HEADS AND DOWNLOAD ALL THE HEADS PARAMETERS
   //ALL THE PARAMETERS ARE AVAILABLE ON THE CONSTANTS STRUCTURE

   //If all head initialized. Jump back

   #TMP_xWriteDoneOS := 0;

   //Check the condition to set the initialization step
       //Only download parameters to the head not initialized and with IP link available
   IF NOT (#ST_xHeadInitialized) AND (#ST_xHeadIPAvail) AND NOT (#tALM.tS.x0) THEN
           #PH_xHeadInit := 1;
       END_IF;

       IF (#PH_xHeadInit) THEN
           IF (#AUX_dActualDownloadPar < "PLANT_CONSTANTS".CONST_rgtHeadPar[#IN_dHeadCycleIndex].dParametersToDownload) THEN

               //No action in progress, ask the execution of the download
               IF (NOT (#ILx2T_Parameter_Read_Write_Instance.q_xWriteDone) AND NOT (#ILx2T_Parameter_Read_Write_Instance.q_xBusy) AND NOT (#ILx2T_Parameter_Read_Write_Instance.q_xError))
                   AND  #ILx2T_Parameter_Read_Write_Instance.i_xParameterWrite = 0 THEN //AND NOT(#AUX_tmWaitWriteParam.Q) THEN
                   //Prepare information for download
                   #TMP_dIndex2Nd := #AUX_dActualDownloadPar;
                   #ILx2T_Parameter_Read_Write_Instance.i_woParameterAddress := INT_TO_WORD("PLANT_CONSTANTS".CONST_rgtHeadPar[#IN_dHeadCycleIndex].rgtAxisParameters[#TMP_dIndex2Nd].iAddress);
                   #ILx2T_Parameter_Read_Write_Instance.i_diWriteParameterValue := "PLANT_CONSTANTS".CONST_rgtHeadPar[#IN_dHeadCycleIndex].rgtAxisParameters[#TMP_dIndex2Nd].dValue;
                   #ILx2T_Parameter_Read_Write_Instance.i_byWriteParameterLength := "PLANT_CONSTANTS".CONST_rgtHeadPar[#IN_dHeadCycleIndex].rgtAxisParameters[#TMP_dIndex2Nd].iLength;

                   #ILx2T_Parameter_Read_Write_Instance.i_xParameterWrite := 1;

               END_IF;

               //Check the result of the execution. If busy wait; if done proceed to the next parameters; if error retry           
               IF (#ILx2T_Parameter_Read_Write_Instance.q_xWriteDone) AND  #ILx2T_Parameter_Read_Write_Instance.i_xParameterWrite = 1 THEN  //AND NOT(#AUX_tmWaitWriteParam.Q) THEN
                   #AUX_dActualDownloadPar := #AUX_dActualDownloadPar + 1;
                   #ILx2T_Parameter_Read_Write_Instance.i_xParameterWrite := 0;

               END_IF;

               //Execution done with error. Retry.... The timeout anomaly will reinitialize the download
               IF (#ILx2T_Parameter_Read_Write_Instance.q_xError) THEN
                   #ILx2T_Parameter_Read_Write_Instance.i_xParameterWrite := 0;
               END_IF;


           ELSE
               //Download parameters done
               #ST_xHeadInitialized := 1;
               #PH_xHeadInit := 0;
               #AUX_dActualDownloadPar := 0;
               #TMP_xWriteDoneOS := 1;
           END_IF;
       ELSE

           #ILx2T_Parameter_Read_Write_Instance.i_xParameterWrite := 0;

       END_IF;

       IF #ST_xBrakeReleaseRequest THEN
           #ILx2T_Parameter_Read_Write_Instance.i_xParameterWrite := 1;
       END_IF;


       IF ((#ST_xHeadInitialized) OR (#ILx2T_Parameter_Read_Write_Instance_Pos.q_xBusy) OR (#ILx2T_Parameter_Read_Write_Instance_Pos.q_xError)
           OR (#ILx2T_Parameter_Read_Write_Instance_Speed.q_xBusy) OR (#ILx2T_Parameter_Read_Write_Instance_Speed.q_xError)) AND NOT(#ST_xBrakeReleaseRequest) THEN
           #ILx2T_Parameter_Read_Write_Instance.i_xParameterWrite := 0;
       END_IF;
END_REGION

REGION Network 26: Call fb read write parameter
   RUNG wire#powerrail
      #ILx2T_Parameter_Read_Write_Instance(i_xParameterRead :=, i_xParameterWrite :=, i_woParameterAddress :=, i_byWriteParameterLength :=, i_diWriteParameterValue :=, ILx2T_Ref := #Axis_Ref, q_xReadValueValid =>, q_xWriteDone =>, q_xError =>, q_xBusy =>, q_diReadParameterValue =>)
   END_RUNG
   // the same network as SCL:
   #ILx2T_Parameter_Read_Write_Instance(ILx2T_Ref := #Axis_Ref);   // "ILx2T_Parameter_Read_Write"
END_REGION

REGION Network 27: Power on motors
   #AUX_tmDriveReadyRetainTimer.TOF(IN := (#ST_xOutputEnable AND (#PH_xHeadHomeSwitch OR #PH_xHeadEndHomeSwitch OR #PH_xHeadPositioning OR #PH_xHeadEndPositioning)) OR ("Z256".ST_xManualModeAccepted AND (#tHMW.tManCmd.xMan_JogForward OR #tHMW.tManCmd.xMan_JogBackward)),
                           PT := T#100MS);
END_REGION

REGION Network 28: Enable drive
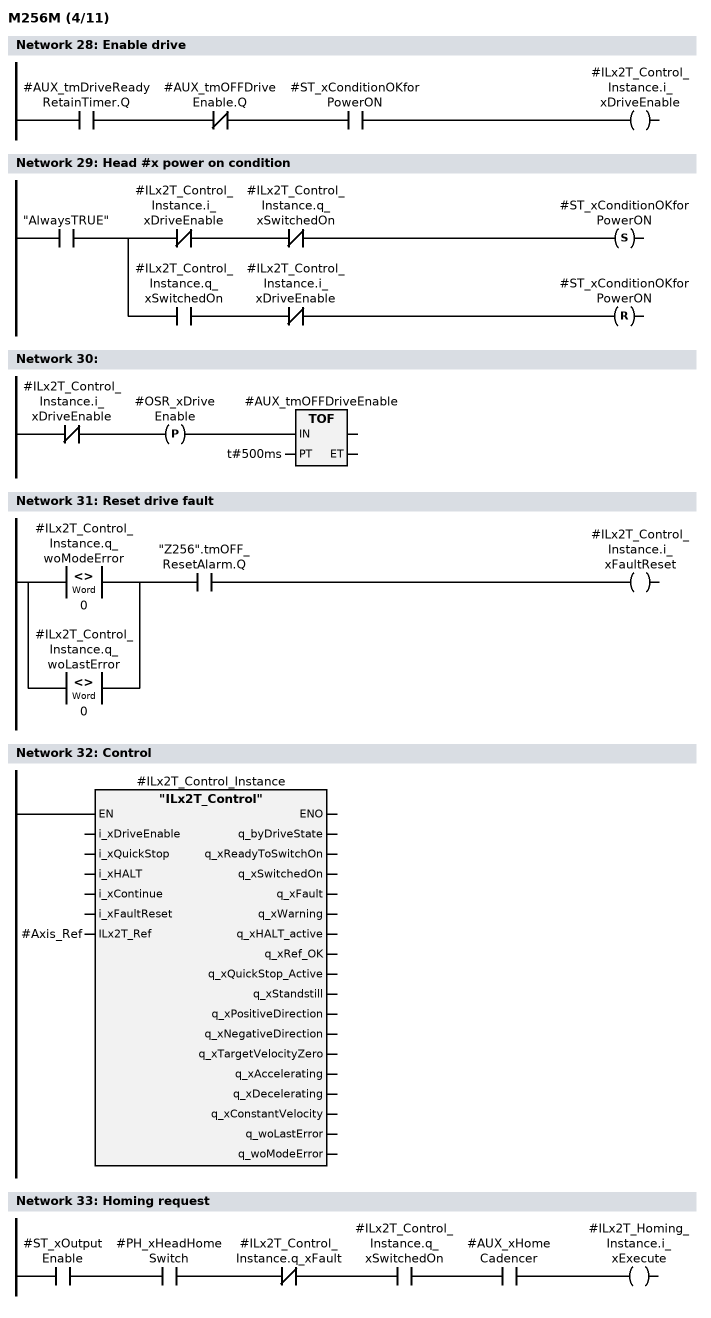
   RUNG wire#powerrail
      Contact( #AUX_tmDriveReadyRetainTimer.Q )
      I_Contact( #AUX_tmOFFDriveEnable.Q )
      Contact( #ST_xConditionOKforPowerON )
      Coil( #ILx2T_Control_Instance.i_xDriveEnable )
   END_RUNG
   // the same network as SCL:
   #ILx2T_Control_Instance.i_xDriveEnable := #AUX_tmDriveReadyRetainTimer.Q AND NOT #AUX_tmOFFDriveEnable.Q AND #ST_xConditionOKforPowerON;
END_REGION

REGION Network 29: Head #x power on condition
   RUNG wire#powerrail
      Contact( "AlwaysTRUE" )
      wire#w1
      I_Contact( #ILx2T_Control_Instance.i_xDriveEnable )
      I_Contact( #ILx2T_Control_Instance.q_xSwitchedOn )
      S_Coil( #ST_xConditionOKforPowerON )
   END_RUNG
   RUNG wire#w1
      Contact( #ILx2T_Control_Instance.q_xSwitchedOn )
      I_Contact( #ILx2T_Control_Instance.i_xDriveEnable )
      R_Coil( #ST_xConditionOKforPowerON )
   END_RUNG
   // the same network as SCL:
   IF "AlwaysTRUE" AND NOT #ILx2T_Control_Instance.i_xDriveEnable AND NOT #ILx2T_Control_Instance.q_xSwitchedOn THEN
       #ST_xConditionOKforPowerON := TRUE;
   END_IF;
   IF "AlwaysTRUE" AND #ILx2T_Control_Instance.q_xSwitchedOn AND NOT #ILx2T_Control_Instance.i_xDriveEnable THEN
       #ST_xConditionOKforPowerON := FALSE;
   END_IF;
END_REGION

REGION Network 30
   #_w1 := NOT #ILx2T_Control_Instance.i_xDriveEnable AND NOT #OSR_xDriveEnable;   // rising edge
   #OSR_xDriveEnable := NOT #ILx2T_Control_Instance.i_xDriveEnable;
   #AUX_tmOFFDriveEnable.TOF(IN := #_w1, PT := t#500ms);
END_REGION

REGION Network 31: Reset drive fault
   RUNG wire#powerrail
      { S7_Templates := "SrcType := Word" } NE_Contact(in1 := #ILx2T_Control_Instance.q_woModeError, in2 := 0)
      wire#w1
      Contact( "Z256".tmOFF_ResetAlarm.Q )
      Coil( #ILx2T_Control_Instance.i_xFaultReset )
   END_RUNG
   RUNG wire#powerrail
      { S7_Templates := "SrcType := Word" } NE_Contact(in1 := #ILx2T_Control_Instance.q_woLastError, in2 := 0)
   END_RUNG wire#w1
   // the same network as SCL:
   #ILx2T_Control_Instance.i_xFaultReset := ((#ILx2T_Control_Instance.q_woModeError <> 0) OR (#ILx2T_Control_Instance.q_woLastError <> 0)) AND "Z256".tmOFF_ResetAlarm.Q;
END_REGION

REGION Network 32: Control
   RUNG wire#powerrail
      #ILx2T_Control_Instance(i_xDriveEnable :=, i_xQuickStop :=, i_xHALT :=, i_xContinue :=, i_xFaultReset :=, ILx2T_Ref := #Axis_Ref, q_byDriveState =>, q_xReadyToSwitchOn =>, q_xSwitchedOn =>, q_xFault =>, q_xWarning =>, q_xHALT_active =>, q_xRef_OK =>, q_xQuickStop_Active =>, q_xStandstill =>, q_xPositiveDirection =>, q_xNegativeDirection =>, q_xTargetVelocityZero =>, q_xAccelerating =>, q_xDecelerating =>, q_xConstantVelocity =>, q_woLastError =>, q_woModeError =>)
   END_RUNG
   // the same network as SCL:
   #ILx2T_Control_Instance(ILx2T_Ref := #Axis_Ref);   // "ILx2T_Control"
END_REGION

REGION Network 33: Homing request
   RUNG wire#powerrail
      Contact( #ST_xOutputEnable )
      Contact( #PH_xHeadHomeSwitch )
      I_Contact( #ILx2T_Control_Instance.q_xFault )
      Contact( #ILx2T_Control_Instance.q_xSwitchedOn )
      Contact( #AUX_xHomeCadencer )
      Coil( #ILx2T_Homing_Instance.i_xExecute )
   END_RUNG
   // the same network as SCL:
   #ILx2T_Homing_Instance.i_xExecute := #ST_xOutputEnable AND #PH_xHeadHomeSwitch AND NOT #ILx2T_Control_Instance.q_xFault AND #ILx2T_Control_Instance.q_xSwitchedOn AND #AUX_xHomeCadencer;
END_REGION

REGION Network 34: Homing